
         O     "DB619_State_MPart".Cycle[1].LastStanbyTimeTool;
         O     "DB110_Interf_Program_M1".Bits.MouldNotReleased;
         =     "DB110_Interf_Program_M1".Bits.LastStandbyTimeTool;
END_REGION

REGION Network 6: Interface signals mixinghead 1 mouldcarrier 1
         A     "DB704_MH_Value".MH_Inerting[1].with_output_without_N2;
         =     "DB614_MH_State".InertingMH[1].Inert_Off_Dry_Shot;

         O     "DB123_MH_IO_Signals".MH[1].IN.MH_Manual_Mode;
         O     "DB123_MH_IO_Signals".MH[1].IN.MH_Auto_Mode;
         AN    "DB824_Error_MH_CP".MH_Control[1].FLT_ShotStopped;
         AN    "DB824_Error_MH_CP".CPiston[1].IPS_defect;
         A     "DB619_State_MPart".Operationmode[1].Auto;
         A     "DB619_State_MPart".Operationmode[1].Active;
         =     #Release_Foaming;
   //------------------------------------------------------------------------------
   //  Freigabe zum automatischen Abruf des Schäumzykluses
   //------------------------------------------------------------------------------
   //-----
         O     "DB005_RS<->Extern".MC_Interface[1].Data_from_MC.Shot_preperation;
         O     "DB005_RS<->Extern".MC_Interface[1].Data_from_MC.Shot_release;
         =     #TempReleasInterface;
   //-----
         O     "DB110_Interf_Program_M1".HM_MC_Fault."01";
         =     "DB123_MH_IO_Signals".MH[1].OUT.MH.K_Fault_MC;
         =     "DB005_RS<->Extern".MC_Interface[1].Data_to_MC.Fault;
   //------------------------------------------------------------------------------
   // Programmno. interface in manual mode
   //------------------------------------------------------------------------------
         L     "DB123_MH_IO_Signals".MH[1].IN.MH_Prog_No_MH;
         A     "DB123_MH_IO_Signals".MH[1].IN.MH_Manual_Mode;
         JC    prnr;
         L     0;
   prnr: T     #Temp_ProgNo_MK1_manual;
   //-----
         A     "DB123_MH_IO_Signals".MH[1].IN.MH_Start;
         A     "DB123_MH_IO_Signals".MH[1].IN.MH_Manual_Mode;
         =     #Start_Zyklus;
   //-----
         O(;
         A     "DB005_RS<->Extern".MC_Interface[1].Data_from_MC.Selected;
         A     "DB123_MH_IO_Signals".MH[1].IN.MH_Stop;
         A     "DB123_MH_IO_Signals".MH[1].IN.MH_Auto_Mode;
         );
         O(;
         A     "DB123_MH_IO_Signals".MH[1].IN.MH_Stop;
         A     "DB123_MH_IO_Signals".MH[1].IN.MH_Manual_Mode;
         );
         =     #Temp_Stop;

   //-----
         CALL  "FC112_IF_SP_MC"
         ( IN_InterfaceNo           := 1,
           IN_PositionFIRST         := "DB110_Interf_Program_M1".FIRST,
           IN_PositionSECOND        := "DB110_Interf_Program_M1".SECOND,
           IN_BCDSwitchPrgrNo_MH    := #Temp_ProgNo_MK1_manual,
           IN_MH_Automatic          := "DB123_MH_IO_Signals".MH[1].IN.MH_Auto_Mode,
           IN_MH_Manual             := "DB123_MH_IO_Signals".MH[1].IN.MH_Manual_Mode,
           IN_Start_MH_Panel        := #Start_Zyklus,  //"DB123_MH_IO_Signals".MH[1].IN.MH_Start
           IN_Stop_MH_Panel         := #Temp_Stop,
           IN_ResetFault            := "DB009_Faults".Faults_Reset_FKT_M1,
           IN_ReleaseSWU            := "DB619_State_MPart".SWU[1].SWU_released."01",
           IN_ReleaseMouldcarrier   := #TempReleasInterface,
           IN_PrgNoSwitchDeselected := "DB123_MH_IO_Signals".MH[1].IN.MH_Auto_Mode,
           IN_ReleaseFoaming        := #Release_Foaming,
           IN_ReleaseCycle          := "DB619_State_MPart".Cycle[1].Release,
           IN_OperationModeAuto     := "DB619_State_MPart".Operationmode[1].Auto,
           IN_OperationModeTest     := "DB619_State_MPart".Operationmode[1].Test,
           IN_LampTest              := "DB619_State_MPart".Operationmode[1].Lamptest,
           IN_CycleRunning          := "DB619_State_MPart".ToolMa[1].StationActive,
           IN_ShotRunning           := "DB619_State_MPart".Cycle[1].ShotRuns,
           IN_LastStandbyTimeCycle  := "DB110_Interf_Program_M1".Bits.LastStandbyTimeTool,
           IN_PulseCycleFinished    := "DB619_State_MPart".Cycle[1].Pulse_ToolFinished,
           OUT_Fault_To_MC          := "DB110_Interf_Program_M1".HM_MC_Fault."01",
           OUT_ShotEnd_To_MC        := "DB110_Interf_Program_M1".HM_MC_Shotend."01",
           OUT_H_MH_Panel           := #H_MH_Panel,  // "DB110_Interf_Program_M1".HM_MC_Lamp."01"
           IO_InterfaceActiveFIFO   := "DB110_Interf_Program_M1".Putin_FIFOlist."01",
           IO_Status                := "DB110_Interf_Program_M1".Status_IF[1],
           IO_Fault                 := "DB825_Error_Interface".Interface_MC[1],
           IO_NewFault              := "DB009_Faults".Faultschanging_M1,
           IO_FaultLevel_1          := "DB009_Faults".Faults_FKT_Grp_1_M1,
           IO_FaultLevel_3          := "DB009_Faults".Faults_FKT_Grp_3_M1
         );
   //-----
   //-
   //- General
   //-
         A     #H_MH_Panel;
         O(;
         A     "DB1900_IF_Robots".State_ABB[1].Output.doIRBInHome;
         A     "DB1900_IF_Robots".State_ABB[1].Output.doIRBinAuto;
         A     "DB1900_IF_Robots".State_ABB[1].Output.doCycleOn;
         AN    "DB1900_IF_Robots".State_ABB[1].Output.doSysError;
         AN    "DB619_State_MPart".Cycle[1].running;
         );
         O(;
         A     "DB1900_IF_Robots".State_ABB[1].Output.doIRBInWaitP;
         A     "DB1900_IF_Robots".State_ABB[1].Output.doInWaitPos;
         );
         AN    "DB619_State_MPart".Operationmode[1].Test;
         O     "DB110_Interf_Program_M1".Test_M01.Spare_0_7;
         =     "DB110_Interf_Program_M1".HM_MC_Lamp."01";
   //----------------------------------------------------------------------------------------
   //     Schnittstelle Presse
   //----------------------------------------------------------------------------------------
         AN    #TempReleasInterface;
         R     "DB005_RS<->Extern".MC_Interface[1].Data_to_MC.Shot_end;
   //
         O     "DB110_Interf_Program_M1".Bits.MouldNotReleased;
         O(;
         A     #TempReleasInterface;
         A     "DB110_Interf_Program_M1".HM_MC_Shotend."01";
         );
         S     "DB005_RS<->Extern".MC_Interface[1].Data_to_MC.Shot_end;
   //
         A     "DB005_RS<->Extern".MC_Interface[1].Data_to_MC.Shot_end;
         =     "DB123_MH_IO_Signals".MH[1].OUT.MH.K_ShotEnd_MC;
   //-----
         A     "DB110_Interf_Program_M1".HM_MC_Fault."01";
         =     "DB005_RS<->Extern".MC_Interface[1].Data_to_MC.Fault;
   //
         A     "DB123_MH_IO_Signals".MH[1].IN.MH_Auto_Mode;
         A     "DB619_State_MPart".Operationmode[1].Auto;
         =     "DB005_RS<->Extern".MC_Interface[1].Data_to_MC.Automatic_mode;
   //
         AN    "DB614_MH_State".MH_Status[1].Switch_Service_ON_OFF;
         =     "DB005_RS<->Extern".MC_Interface[1].Data_to_MC.Service_mode;
   //
         A     "DB619_State_MPart".Cycle[1].ShotRuns;
         =     "DB005_RS<->Extern".MC_Interface[1].Data_to_MC.Shot_runs;
   //
         O     "DB1900_IF_Robots".State_ABB[1].Output.doIRBInHome;
         O     "DB1900_IF_Robots".State_ABB[1].Output.doSafetyArea_1;
         =     "DB005_RS<->Extern".MC_Interface[1].Data_to_MC.Robot_out_of_MC;
   //
         A     "DB005_RS<->Extern".MC_Interface[1].Data_from_MC.Com_control;
         =     "DB005_RS<->Extern".MC_Interface[1].Data_to_MC.Com_Control;
   //
         L     "DB005_RS<->Extern".MC_Interface[1].Data_from_MC.Toolcode;
         T     "DB005_RS<->Extern".MC_Interface[1].Data_to_MC.Toolcode;
   //-----
         A     "DB009_Faults".Faults_Reset_FKT_M1;
         R     "DB825_Error_Interface".Interface_MC[1].FLT_Communication;

         L     s5t#5s;
         AN    "DB005_RS<->Extern".MC_Interface[1].Data_from_MC.Com_control;
         SE    "TIM_FRA_WDG1";

         AN    "TIM_FRA_WDG1";
         AN    "DB825_Error_Interface".Interface_MC[1].FLT_Communication;
         CLR;
         S     "DB825_Error_Interface".Interface_MC[1].FLT_Communication;

   // load number to tool alloc
         AN    "DB790_PlantParameter".Bit.ProgrammNofromInterface;
         JC    NoToolNoFromIF01;

         CALL  "FC5_Check_allocAutoMode"
         ( ToolcodeNo := "DB005_RS<->Extern".MC_Interface[1].Data_from_MC.Toolcode,
           ToolAlloc  := "DB940_Tool_alloc_automatic".Alloc_stationTool[1]
         );

   NoToolNoFromIF01:NOP   0;
END_REGION

REGION Network 7: Interface signals mixinghead 2 mouldcarrier 2
         A     "DB704_MH_Value".MH_Inerting[1].with_output_without_N2;
         =     "DB614_MH_State".InertingMH[1].Inert_Off_Dry_Shot;

         O     "DB123_MH_IO_Signals".MH[1].IN.MH_Manual_Mode;
         O     "DB123_MH_IO_Signals".MH[1].IN.MH_Auto_Mode;
         AN    "DB824_Error_MH_CP".MH_Control[1].FLT_ShotStopped;
         AN    "DB824_Error_MH_CP".CPiston[1].IPS_defect;
         A     "DB619_State_MPart".Operationmode[1].Auto;
         A     "DB619_State_MPart".Operationmode[1].Active;
         =     #Release_Foaming;
   //------------------------------------------------------------------------------
   //  Freigabe zum automatischen Abruf des Schäumzykluses
   //------------------------------------------------------------------------------
   //-----
         O     "DB005_RS<->Extern".MC_Interface[2].Data_from_MC.Shot_preperation;
         O     "DB005_RS<->Extern".MC_Interface[2].Data_from_MC.Shot_release;
         =     #TempReleasInterface;
   //-----
         O     "DB110_Interf_Program_M1".HM_MC_Fault."02";
         =     "DB005_RS<->Extern".MC_Interface[2].Data_to_MC.Fault;
   //-----
         A     "DB123_MH_IO_Signals".MH[1].IN.MH_Start;
         A     "DB123_MH_IO_Signals".MH[1].IN.MH_Manual_Mode;
         =     #Start_Zyklus;
   //-----
         A     "DB005_RS<->Extern".MC_Interface[2].Data_from_MC.Selected;
         A     "DB123_MH_IO_Signals".MH[1].IN.MH_Stop;
         =     #Temp_Stop;
   //-----
         CALL  "FC112_IF_SP_MC"
         ( IN_InterfaceNo           := 2,
           IN_PositionFIRST         := "DB110_Interf_Program_M1".FIRST,
           IN_PositionSECOND        := "DB110_Interf_Program_M1".SECOND,
           IN_BCDSwitchPrgrNo_MH    := 0,
           IN_MH_Automatic          := "DB123_MH_IO_Signals".MH[1].IN.MH_Auto_Mode,
           IN_MH_Manual             := false,
           IN_Start_MH_Panel        := #Start_Zyklus,
           IN_Stop_MH_Panel         := #Temp_Stop,
           IN_ResetFault            := "DB009_Faults".Faults_Reset_FKT_M1,
           IN_ReleaseSWU            := "DB619_State_MPart".SWU[1].SWU_released."01",
           IN_ReleaseMouldcarrier   := #TempReleasInterface,
           IN_PrgNoSwitchDeselected := "DB123_MH_IO_Signals".MH[1].IN.MH_Auto_Mode,
           IN_ReleaseFoaming        := #Release_Foaming,
           IN_ReleaseCycle          := "DB619_State_MPart".Cycle[1].Release,
           IN_OperationModeAuto     := "DB619_State_MPart".Operationmode[1].Auto,
           IN_OperationModeTest     := "DB619_State_MPart".Operationmode[1].Test,
           IN_LampTest              := "DB619_State_MPart".Operationmode[1].Lamptest,
           IN_CycleRunning          := "DB619_State_MPart".ToolMa[1].StationActive,
           IN_ShotRunning           := "DB619_State_MPart".Cycle[1].ShotRuns,
           IN_LastStandbyTimeCycle  := "DB110_Interf_Program_M1".Bits.LastStandbyTimeTool,
           IN_PulseCycleFinished    := "DB619_State_MPart".Cycle[1].Pulse_ToolFinished,
           OUT_Fault_To_MC          := "DB110_Interf_Program_M1".HM_MC_Fault."02",
           OUT_ShotEnd_To_MC        := "DB110_Interf_Program_M1".HM_MC_Shotend."02",
           OUT_H_MH_Panel           := #H_MH_Panel,  // "DB110_Interf_Program_M1".HM_MC_Lamp."02"
           IO_InterfaceActiveFIFO   := "DB110_Interf_Program_M1".Putin_FIFOlist."02",
           IO_Status                := "DB110_Interf_Program_M1".Status_IF[2],
           IO_Fault                 := "DB825_Error_Interface".Interface_MC[2],
           IO_NewFault              := "DB009_Faults".Faultschanging_M1,
           IO_FaultLevel_1          := "DB009_Faults".Faults_FKT_Grp_1_M1,
           IO_FaultLevel_3          := "DB009_Faults".Faults_FKT_Grp_3_M1
         );
   //-----
   //-
   //- General
   //-
         A     #H_MH_Panel;
         O(;
         A     "DB1900_IF_Robots".State_ABB[1].Output.doIRBInHome;
         A     "DB1900_IF_Robots".State_ABB[1].Output.doIRBinAuto;
         A     "DB1900_IF_Robots".State_ABB[1].Output.doCycleOn;
         AN    "DB1900_IF_Robots".State_ABB[1].Output.doSysError;
         AN    "DB619_State_MPart".Cycle[1].running;
         );
         O(;
         A     "DB1900_IF_Robots".State_ABB[1].Output.doIRBInWaitP;
         A     "DB1900_IF_Robots".State_ABB[1].Output.doInWaitPos;
         );
         =     "DB110_Interf_Program_M1".HM_MC_Lamp."02";
   //----------------------------------------------------------------------------------------
   //     Schnittstelle Presse
   //----------------------------------------------------------------------------------------
         AN    #TempReleasInterface;
         R     "DB005_RS<->Extern".MC_Interface[2].Data_to_MC.Shot_end;
   //
         O     "DB110_Interf_Program_M1".Bits.MouldNotReleased;
         O(;
         A     #TempReleasInterface;
         A     "DB110_Interf_Program_M1".HM_MC_Shotend."02";
         );
         S     "DB005_RS<->Extern".MC_Interface[2].Data_to_MC.Shot_end;
   //-----
         A     "DB110_Interf_Program_M1".HM_MC_Fault."02";
         =     "DB005_RS<->Extern".MC_Interface[2].Data_to_MC.Fault;
   //
         A     "DB123_MH_IO_Signals".MH[1].IN.MH_Auto_Mode;
         A     "DB619_State_MPart".Operationmode[1].Auto;
         =     "DB005_RS<->Extern".MC_Interface[2].Data_to_MC.Automatic_mode;
   //
         AN    "DB614_MH_State".MH_Status[1].Switch_Service_ON_OFF;
         =     "DB005_RS<->Extern".MC_Interface[2].Data_to_MC.Service_mode;
   //
         A     "DB619_State_MPart".Cycle[1].ShotRuns;
         =     "DB005_RS<->Extern".MC_Interface[2].Data_to_MC.Shot_runs;
   //
         O     "DB1900_IF_Robots".State_ABB[1].Output.doIRBInHome;
         O     "DB1900_IF_Robots".State_ABB[1].Output.doSafetyArea_2;
         =     "DB005_RS<->Extern".MC_Interface[2].Data_to_MC.Robot_out_of_MC;
   //
         A     "DB005_RS<->Extern".MC_Interface[2].Data_from_MC.Com_control;
         =     "DB005_RS<->Extern".MC_Interface[2].Data_to_MC.Com_Control;
   //
         L     "DB005_RS<->Extern".MC_Interface[2].Data_from_MC.Toolcode;
         T     "DB005_RS<->Extern".MC_Interface[2].Data_to_MC.Toolcode;
   //-----
         A     "DB009_Faults".Faults_Reset_FKT_M1;
         R     "DB825_Error_Interface".Interface_MC[2].FLT_Communication;

         L     s5t#5s;
         AN    "DB005_RS<->Extern".MC_Interface[2].Data_from_MC.Com_control;
         SE    "TIM_FRA_WDG2";

         AN    "TIM_FRA_WDG2";
         AN    "DB825_Error_Interface".Interface_MC[2].FLT_Communication;
         CLR;
         S     "DB825_Error_Interface".Interface_MC[2].FLT_Communication;

   // load number to tool alloc
         AN    "DB790_PlantParameter".Bit.ProgrammNofromInterface;
         JC    NoToolNoFromIF02;

         CALL  "FC5_Check_allocAutoMode"
         ( ToolcodeNo := "DB005_RS<->Extern".MC_Interface[2].Data_from_MC.Toolcode,
           ToolAlloc  := "DB940_Tool_alloc_automatic".Alloc_stationTool[2]
         );

   NoToolNoFromIF02:NOP   0;
END_REGION

REGION Network 8: Interface signals mixinghead 3 mouldcarrier 3
         A     "DB704_MH_Value".MH_Inerting[1].with_output_without_N2;
         =     "DB614_MH_State".InertingMH[1].Inert_Off_Dry_Shot;

         O     "DB123_MH_IO_Signals".MH[1].IN.MH_Manual_Mode;
         O     "DB123_MH_IO_Signals".MH[1].IN.MH_Auto_Mode;
         AN    "DB824_Error_MH_CP".MH_Control[1].FLT_ShotStopped;
         AN    "DB824_Error_MH_CP".CPiston[1].IPS_defect;
         A     "DB619_State_MPart".Operationmode[1].Auto;
         A     "DB619_State_MPart".Operationmode[1].Active;
         =     #Release_Foaming;
   //------------------------------------------------------------------------------
   //  Freigabe zum automatischen Abruf des Schäumzykluses
   //------------------------------------------------------------------------------
   //-----
         O     "DB005_RS<->Extern".MC_Interface[3].Data_from_MC.Shot_preperation;
         O     "DB005_RS<->Extern".MC_Interface[3].Data_from_MC.Shot_release;
         =     #TempReleasInterface;
   //-----
         O     "DB110_Interf_Program_M1".HM_MC_Fault."03";
         =     "DB005_RS<->Extern".MC_Interface[3].Data_to_MC.Fault;
   //-----
         A     "DB123_MH_IO_Signals".MH[1].IN.MH_Start;
         A     "DB123_MH_IO_Signals".MH[1].IN.MH_Manual_Mode;
         =     #Start_Zyklus;
   //-----
         A     "DB005_RS<->Extern".MC_Interface[3].Data_from_MC.Selected;
         A     "DB123_MH_IO_Signals".MH[1].IN.MH_Stop;
         =     #Temp_Stop;
   //-----
         CALL  "FC112_IF_SP_MC"
         ( IN_InterfaceNo           := 3,
           IN_PositionFIRST         := "DB110_Interf_Program_M1".FIRST,
           IN_PositionSECOND        := "DB110_Interf_Program_M1".SECOND,
           IN_BCDSwitchPrgrNo_MH    := 0,
           IN_MH_Automatic          := "DB123_MH_IO_Signals".MH[1].IN.MH_Auto_Mode,
           IN_MH_Manual             := false,
           IN_Start_MH_Panel        := #Start_Zyklus,
           IN_Stop_MH_Panel         := #Temp_Stop,
           IN_ResetFault            := "DB009_Faults".Faults_Reset_FKT_M1,
           IN_ReleaseSWU            := "DB619_State_MPart".SWU[1].SWU_released."01",
           IN_ReleaseMouldcarrier   := #TempReleasInterface,
           IN_PrgNoSwitchDeselected := "DB123_MH_IO_Signals".MH[1].IN.MH_Auto_Mode,
           IN_ReleaseFoaming        := #Release_Foaming,
           IN_ReleaseCycle          := "DB619_State_MPart".Cycle[1].Release,
           IN_OperationModeAuto     := "DB619_State_MPart".Operationmode[1].Auto,
           IN_OperationModeTest     := "DB619_State_MPart".Operationmode[1].Test,
           IN_LampTest              := "DB619_State_MPart".Operationmode[1].Lamptest,
           IN_CycleRunning          := "DB619_State_MPart".ToolMa[1].StationActive,
           IN_ShotRunning           := "DB619_State_MPart".Cycle[1].ShotRuns,
           IN_LastStandbyTimeCycle  := "DB110_Interf_Program_M1".Bits.LastStandbyTimeTool,
           IN_PulseCycleFinished    := "DB619_State_MPart".Cycle[1].Pulse_ToolFinished,
           OUT_Fault_To_MC          := "DB110_Interf_Program_M1".HM_MC_Fault."03",
           OUT_ShotEnd_To_MC        := "DB110_Interf_Program_M1".HM_MC_Shotend."03",
           OUT_H_MH_Panel           := #H_MH_Panel,  // "DB110_Interf_Program_M1".HM_MC_Lamp."03"
           IO_InterfaceActiveFIFO   := "DB110_Interf_Program_M1".Putin_FIFOlist."03",
           IO_Status                := "DB110_Interf_Program_M1".Status_IF[3],
           IO_Fault                 := "DB825_Error_Interface".Interface_MC[3],
           IO_NewFault              := "DB009_Faults".Faultschanging_M1,
           IO_FaultLevel_1          := "DB009_Faults".Faults_FKT_Grp_1_M1,
           IO_FaultLevel_3          := "DB009_Faults".Faults_FKT_Grp_3_M1
         );
   //-----
   //-
   //- General
   //-
         A     #H_MH_Panel;
         O(;
         A     "DB1900_IF_Robots".State_ABB[1].Output.doIRBInHome;
         A     "DB1900_IF_Robots".State_ABB[1].Output.doIRBinAuto;
         A     "DB1900_IF_Robots".State_ABB[1].Output.doCycleOn;
         AN    "DB1900_IF_Robots".State_ABB[1].Output.doSysError;
         AN    "DB619_State_MPart".Cycle[1].running;
         );
         O(;
         A     "DB1900_IF_Robots".State_ABB[1].Output.doIRBInWaitP;
         A     "DB1900_IF_Robots".State_ABB[1].Output.doInWaitPos;
         );
         =     "DB110_Interf_Program_M1".HM_MC_Lamp."03";
   //----------------------------------------------------------------------------------------
   //     Schnittstelle Presse
   //----------------------------------------------------------------------------------------
         AN    #TempReleasInterface;
         R     "DB005_RS<->Extern".MC_Interface[3].Data_to_MC.Shot_end;
   //
         O     "DB110_Interf_Program_M1".Bits.MouldNotReleased;
         O(;
         A     #TempReleasInterface;
         A     "DB110_Interf_Program_M1".HM_MC_Shotend."03";
         );
         S     "DB005_RS<->Extern".MC_Interface[3].Data_to_MC.Shot_end;
   //-----
         A     "DB110_Interf_Program_M1".HM_MC_Fault."03";
         =     "DB005_RS<->Extern".MC_Interface[3].Data_to_MC.Fault;
   //
         A     "DB123_MH_IO_Signals".MH[1].IN.MH_Auto_Mode;
         A     "DB619_State_MPart".Operationmode[1].Auto;
         =     "DB005_RS<->Extern".MC_Interface[3].Data_to_MC.Automatic_mode;
   //
         AN    "DB614_MH_State".MH_Status[1].Switch_Service_ON_OFF;
         =     "DB005_RS<->Extern".MC_Interface[3].Data_to_MC.Service_mode;
   //
         A     "DB619_State_MPart".Cycle[1].ShotRuns;
         =     "DB005_RS<->Extern".MC_Interface[3].Data_to_MC.Shot_runs;
   //
         O     "DB1900_IF_Robots".State_ABB[1].Output.doIRBInHome;
         O     "DB1900_IF_Robots".State_ABB[1].Output.doSafetyArea_3;
         =     "DB005_RS<->Extern".MC_Interface[3].Data_to_MC.Robot_out_of_MC;
   //
         A     "DB005_RS<->Extern".MC_Interface[3].Data_from_MC.Com_control;
         =     "DB005_RS<->Extern".MC_Interface[3].Data_to_MC.Com_Control;
   //
         L     "DB005_RS<->Extern".MC_Interface[3].Data_from_MC.Toolcode;
         T     "DB005_RS<->Extern".MC_Interface[3].Data_to_MC.Toolcode;
   //-----
         A     "DB009_Faults".Faults_Reset_FKT_M1;
         R     "DB825_Error_Interface".Interface_MC[3].FLT_Communication;

         L     s5t#5s;
         AN    "DB005_RS<->Extern".MC_Interface[3].Data_from_MC.Com_control;
         SE    "TIM_FRA_WDG3";

         AN    "TIM_FRA_WDG3";
         A     "With_MC03";
         AN    "DB825_Error_Interface".Interface_MC[3].FLT_Communication;
         S     "DB825_Error_Interface".Interface_MC[3].FLT_Communication;

   // load number to tool alloc
         AN    "DB790_PlantParameter".Bit.ProgrammNofromInterface;
         JC    NoToolNoFromIF03;

         CALL  "FC5_Check_allocAutoMode"
         ( ToolcodeNo := "DB005_RS<->Extern".MC_Interface[3].Data_from_MC.Toolcode,
           ToolAlloc  := "DB940_Tool_alloc_automatic".Alloc_stationTool[3]
         );

   NoToolNoFromIF03:NOP   0;
END_REGION

REGION Network 9: Interface signals mixinghead 4 mouldcarrier 4
         A     "DB704_MH_Value".MH_Inerting[1].with_output_without_N2;
         =     "DB614_MH_State".InertingMH[1].Inert_Off_Dry_Shot;

         O     "DB123_MH_IO_Signals".MH[1].IN.MH_Manual_Mode;
         O     "DB123_MH_IO_Signals".MH[1].IN.MH_Auto_Mode;
         AN    "DB824_Error_MH_CP".MH_Control[1].FLT_ShotStopped;
         AN    "DB824_Error_MH_CP".CPiston[1].IPS_defect;
         A     "DB619_State_MPart".Operationmode[1].Auto;
         A     "DB619_State_MPart".Operationmode[1].Active;
         =     #Release_Foaming;
   //------------------------------------------------------------------------------
   //  Freigabe zum automatischen Abruf des Schäumzykluses
   //------------------------------------------------------------------------------
   //-----
         O     "DB005_RS<->Extern".MC_Interface[4].Data_from_MC.Shot_preperation;
         O     "DB005_RS<->Extern".MC_Interface[4].Data_from_MC.Shot_release;
         =     #TempReleasInterface;
   //-----
         O     "DB110_Interf_Program_M1".HM_MC_Fault."04";
         =     "DB005_RS<->Extern".MC_Interface[4].Data_to_MC.Fault;
   //-----
         A     "DB123_MH_IO_Signals".MH[1].IN.MH_Start;
         A     "DB123_MH_IO_Signals".MH[1].IN.MH_Manual_Mode;
         =     #Start_Zyklus;
   //-----
         A     "DB005_RS<->Extern".MC_Interface[4].Data_from_MC.Selected;
         A     "DB123_MH_IO_Signals".MH[1].IN.MH_Stop;
         =     #Temp_Stop;
   //-----
         CALL  "FC112_IF_SP_MC"
         ( IN_InterfaceNo           := 4,
           IN_PositionFIRST         := "DB110_Interf_Program_M1".FIRST,
           IN_PositionSECOND        := "DB110_Interf_Program_M1".SECOND,
           IN_BCDSwitchPrgrNo_MH    := 0,
           IN_MH_Automatic          := "DB123_MH_IO_Signals".MH[1].IN.MH_Auto_Mode,
           IN_MH_Manual             := false,
           IN_Start_MH_Panel        := #Start_Zyklus,
           IN_Stop_MH_Panel         := #Temp_Stop,
           IN_ResetFault            := "DB009_Faults".Faults_Reset_FKT_M1,
           IN_ReleaseSWU            := "DB619_State_MPart".SWU[1].SWU_released."01",
           IN_ReleaseMouldcarrier   := #TempReleasInterface,
           IN_PrgNoSwitchDeselected := "DB123_MH_IO_Signals".MH[1].IN.MH_Auto_Mode,
           IN_ReleaseFoaming        := #Release_Foaming,
           IN_ReleaseCycle          := "DB619_State_MPart".Cycle[1].Release,
           IN_OperationModeAuto     := "DB619_State_MPart".Operationmode[1].Auto,
           IN_OperationModeTest     := "DB619_State_MPart".Operationmode[1].Test,
           IN_LampTest              := "DB619_State_MPart".Operationmode[1].Lamptest,
           IN_CycleRunning          := "DB619_State_MPart".ToolMa[1].StationActive,
           IN_ShotRunning           := "DB619_State_MPart".Cycle[1].ShotRuns,
           IN_LastStandbyTimeCycle  := "DB110_Interf_Program_M1".Bits.LastStandbyTimeTool,
           IN_PulseCycleFinished    := "DB619_State_MPart".Cycle[1].Pulse_ToolFinished,
           OUT_Fault_To_MC          := "DB110_Interf_Program_M1".HM_MC_Fault."04",
           OUT_ShotEnd_To_MC        := "DB110_Interf_Program_M1".HM_MC_Shotend."04",
           OUT_H_MH_Panel           := #H_MH_Panel,  // "DB110_Interf_Program_M1".HM_MC_Lamp."04"
           IO_InterfaceActiveFIFO   := "DB110_Interf_Program_M1".Putin_FIFOlist."04",
           IO_Status                := "DB110_Interf_Program_M1".Status_IF[4],
           IO_Fault                 := "DB825_Error_Interface".Interface_MC[4],
           IO_NewFault              := "DB009_Faults".Faultschanging_M1,
           IO_FaultLevel_1          := "DB009_Faults".Faults_FKT_Grp_1_M1,
           IO_FaultLevel_3          := "DB009_Faults".Faults_FKT_Grp_3_M1
         );
   //-----
   //-
   //- General
   //-
         A     #H_MH_Panel;
         O(;
         A     "DB1900_IF_Robots".State_ABB[1].Output.doIRBInHome;
         A     "DB1900_IF_Robots".State_ABB[1].Output.doIRBinAuto;
         A     "DB1900_IF_Robots".State_ABB[1].Output.doCycleOn;
         AN    "DB1900_IF_Robots".State_ABB[1].Output.doSysError;
         AN    "DB619_State_MPart".Cycle[1].running;
         );
         O(;
         A     "DB1900_IF_Robots".State_ABB[1].Output.doIRBInWaitP;
         A     "DB1900_IF_Robots".State_ABB[1].Output.doInWaitPos;
         );
         =     "DB110_Interf_Program_M1".HM_MC_Lamp."04";
   //----------------------------------------------------------------------------------------
   //     Schnittstelle Presse
   //----------------------------------------------------------------------------------------
         AN    #TempReleasInterface;
         R     "DB005_RS<->Extern".MC_Interface[4].Data_to_MC.Shot_end;
   //
         O     "DB110_Interf_Program_M1".Bits.MouldNotReleased;
         O(;
         A     #TempReleasInterface;
         A     "DB110_Interf_Program_M1".HM_MC_Shotend."04";
         );
         S     "DB005_RS<->Extern".MC_Interface[4].Data_to_MC.Shot_end;
   //-----
         A     "DB110_Interf_Program_M1".HM_MC_Fault."04";
         =     "DB005_RS<->Extern".MC_Interface[4].Data_to_MC.Fault;
   //
         A     "DB123_MH_IO_Signals".MH[1].IN.MH_Auto_Mode;
         A     "DB619_State_MPart".Operationmode[1].Auto;
         =     "DB005_RS<->Extern".MC_Interface[4].Data_to_MC.Automatic_mode;
   //
         AN    "DB614_MH_State".MH_Status[1].Switch_Service_ON_OFF;
         =     "DB005_RS<->Extern".MC_Interface[4].Data_to_MC.Service_mode;
   //
         A     "DB619_State_MPart".Cycle[1].ShotRuns;
         =     "DB005_RS<->Extern".MC_Interface[4].Data_to_MC.Shot_runs;
   //
         O     "DB1900_IF_Robots".State_ABB[1].Output.doIRBInHome;
         O     "DB1900_IF_Robots".State_ABB[1].Output.doSafetyArea_4;
         =     "DB005_RS<->Extern".MC_Interface[4].Data_to_MC.Robot_out_of_MC;
   //
         A     "DB005_RS<->Extern".MC_Interface[4].Data_from_MC.Com_control;
         =     "DB005_RS<->Extern".MC_Interface[4].Data_to_MC.Com_Control;
   //
         L     "DB005_RS<->Extern".MC_Interface[4].Data_from_MC.Toolcode;
         T     "DB005_RS<->Extern".MC_Interface[4].Data_to_MC.Toolcode;
   //-----
         A     "DB009_Faults".Faults_Reset_FKT_M1;
         R     "DB825_Error_Interface".Interface_MC[4].FLT_Communication;

         L     s5t#5s;
         AN    "DB005_RS<->Extern".MC_Interface[4].Data_from_MC.Com_control;
         SE    "TIM_FRA_WDG4";

         AN    "TIM_FRA_WDG4";
         A     "With_MC04";
         AN    "DB825_Error_Interface".Interface_MC[4].FLT_Communication;
         S     "DB825_Error_Interface".Interface_MC[4].FLT_Communication;

   // load number to tool alloc
         AN    "DB790_PlantParameter".Bit.ProgrammNofromInterface;
         JC    NoToolNoFromIF04;

         CALL  "FC5_Check_allocAutoMode"
         ( ToolcodeNo := "DB005_RS<->Extern".MC_Interface[4].Data_from_MC.Toolcode,
           ToolAlloc  := "DB940_Tool_alloc_automatic".Alloc_stationTool[4]
         );

   NoToolNoFromIF04:NOP   0;
END_REGION

REGION Network 10: Test with test valves
   //     CALL  "FC115_Testen"
   //         IN_Betriebsart_Testen   :="DB619_State_MPart".Operationmode[1].Test
   //         IN_Betriebsart_Betrieb  :="DB619_State_MPart".Operationmode[1].Operation
   //         IN_Lampentest           :="DB619_State_MPart".Operationmode[1].Lamptest
   //         IN_Start_Testen_K1      :="T_Start_Test_C1"
   //         IN_Start_Testen_K2      :="T_Start_Test_C2"
   //         IN_Start_Testen_K3      :=FALSE
   //         IN_Start_Testen_K4      :=FALSE
   //         IN_Stop_Testen          :="T_Stop_Test"
   //         IN_Stoerung_Gruppe_1    :="DB009_Faults".Faults_FKT_Grp_1_M1
   //         IN_Zyklus_Freigabe      :="DB619_State_MPart".Cycle[1].Release
   //         IN_Zyklus_laeuft        :="DB619_State_MPart".ToolMa[1].StationActive
   //         IN_Zyklus_Schuss_laeuft :="DB619_State_MPart".Cycle[1].ShotRuns
   //         IN_Imp_Zyklus_Ende      :="DB619_State_MPart".Cycle[1].Pulse_ToolFinished
   //         IN_Zyklus_KLZ2_u_ff     :="DB619_State_MPart".Cycle[1].LastStanbyTimeTool
   //         OUT_H_Testen_K1         :="H_Test_C1"
   //         OUT_H_Testen_K2         :="H_Test_C2"
   //         OUT_H_Testen_K3         :=#Dummy
   //         OUT_H_Testen_K4         :=#Dummy
   //         OUT_V_Testen_K1         :="V_Test_C1"
   //         OUT_V_Testen_K2         :="V_Test_C2"
   //         OUT_V_Testen_K3         :=#Dummy
   //         OUT_V_Testen_K4         :=#Dummy
   //         IO_Status               :="DB110_Interf_Program_M1".Test_M01
   //
END_REGION

REGION Network 11: LED mixing head panel
   //-----
         A     "DB110_Interf_Program_M1".HM_MC_Lamp."01";
         O;
         A     "DB110_Interf_Program_M1".Status_IF[2].IF_is_on_1_Position;
         A     "DB110_Interf_Program_M1".HM_MC_Lamp."02";
         O;
         A     "DB110_Interf_Program_M1".Status_IF[3].IF_is_on_1_Position;
         A     "DB110_Interf_Program_M1".HM_MC_Lamp."03";
         O;
         A     "DB110_Interf_Program_M1".Status_IF[4].IF_is_on_1_Position;
         A     "DB110_Interf_Program_M1".HM_MC_Lamp."04";
         O;
         A     "DB110_Interf_Program_M1".Status_IF[5].IF_is_on_1_Position;
         A     "DB110_Interf_Program_M1".HM_MC_Lamp."05";
         =     "DB123_MH_IO_Signals".MH[1].OUT.MH.H_Rel_Foaming_MH;
END_REGION

REGION Network 12: Start cycle
         A     "DB1900_IF_Robots".State_Robots[1].ReadyForStartCycle;
         A     "DB123_MH_IO_Signals".MH[1].IN.MH_Auto_Mode;
         O     "DB123_MH_IO_Signals".MH[1].IN.MH_Manual_Mode;
         A(;
         O     "DB110_Interf_Program_M1".Status_IF[1].Start_to_Cycle;
         O     "DB110_Interf_Program_M1".Status_IF[2].Start_to_Cycle;
         O     "DB110_Interf_Program_M1".Status_IF[3].Start_to_Cycle;
         O     "DB110_Interf_Program_M1".Status_IF[4].Start_to_Cycle;
         O     "DB110_Interf_Program_M1".Status_IF[5].Start_to_Cycle;
         O     "DB110_Interf_Program_M1".Status_IF[6].Start_to_Cycle;
         O     "DB110_Interf_Program_M1".Status_IF[7].Start_to_Cycle;
         O     "DB110_Interf_Program_M1".Status_IF[8].Start_to_Cycle;
         O     "DB110_Interf_Program_M1".Status_IF[9].Start_to_Cycle;
         O     "DB110_Interf_Program_M1".Status_IF[10].Start_to_Cycle;
         );
         O     "DB110_Interf_Program_M1".Test_M01.Start_to_Cycle;
         =     #Start_Zyklus;
END_REGION

REGION Network 13: Stop cycle
         O     "DB110_Interf_Program_M1".Status_IF[1].Stop_to_Cycle;
         O     "DB110_Interf_Program_M1".Status_IF[2].Stop_to_Cycle;
         O     "DB110_Interf_Program_M1".Status_IF[3].Stop_to_Cycle;
         O     "DB110_Interf_Program_M1".Status_IF[4].Stop_to_Cycle;
         O     "DB110_Interf_Program_M1".Status_IF[5].Stop_to_Cycle;
         O     "DB110_Interf_Program_M1".Status_IF[6].Stop_to_Cycle;
         O     "DB110_Interf_Program_M1".Status_IF[7].Stop_to_Cycle;
         O     "DB110_Interf_Program_M1".Status_IF[8].Stop_to_Cycle;
         O     "DB110_Interf_Program_M1".Status_IF[9].Stop_to_Cycle;
         O     "DB110_Interf_Program_M1".Status_IF[10].Stop_to_Cycle;
         O     "DB110_Interf_Program_M1".Test_M01.Stop_to_Cycle;
         =     "DB110_Interf_Program_M1".Bits.Stop_Cycle;
         =     "DB619_State_MPart".ToolMa[1].StopCycle;
END_REGION

REGION Network 14: Station number (Program number) to select mould no. ->FB930
         A     #Start_Zyklus;
         AN    "DB619_State_MPart".ToolMa[1].StopCycle;
         JCN   GOON;
   ///----------
         A     "DB619_State_MPart".Operationmode[1].Test;
         JC    Test;
   ///----------
         AN    "DB110_Interf_Program_M1".Status_IF[1].IF_is_on_1_Position;
         JC    SS_2;
   ///----------
         A     "DB123_MH_IO_Signals".MH[1].IN.MH_Auto_Mode;
         JC    SS1A;
   ///----------
         L     #Temp_ProgNo_MK1_manual;
         L     "DB704_MH_Value".Mixinghead[1].pRrgNumberManual;
         +I;
         T     "DB110_Interf_Program_M1".Program_No_01;
         JU    ENDE;
   ///----------
   SS1A: NOP   0;
         AN    "DB005_RS<->Extern".MC_Interface[1].Data_from_MC.Shot_preperation;
         AN    "DB005_RS<->Extern".MC_Interface[1].Data_from_MC.Shot_release;
         ON    "DB619_State_MPart".SWU[1].SWU_released."01";
         JC    ENDE;
   ///----------
         L     1;
         T     "DB110_Interf_Program_M1".Program_No_01;

         L     1;
         T     "DB110_Interf_Program_M1".MixingHeadNo;
         T     "DB110_Interf_Program_M1".Robot_01.MC_Place_Number;

         L     "DB005_RS<->Extern".MC_Interface[1].Data_from_MC.Angle_frame_foaming_pos;
         L     7.0;
         <=R;
         L     1;  //      L     "DB005_RS<->Extern".MC_Interface[1].Data_from_MC.Toolcode
         JC    ProRob01;
         L     1;  // L     "DB005_RS<->Extern".MC_Interface[1].Data_from_MC.Toolcode
         L     100;
         +I;
   ProRob01:T     "DB110_Interf_Program_M1".Robot_01.Robot_ProgNo_Mould_1;
         JU    ENDE;
   ///----------
   SS_2: NOP   0;
         AN    "DB110_Interf_Program_M1".Status_IF[2].IF_is_on_1_Position;
         JC    SS_3;
         A     "DB123_MH_IO_Signals".MH[1].IN.MH_Auto_Mode;
         JC    SS2A;
   ///----------
         L     0;
         T     "DB110_Interf_Program_M1".Program_No_01;
         JU    ENDE;
   ///----------
   SS2A: NOP   0;
         AN    "DB005_RS<->Extern".MC_Interface[2].Data_from_MC.Shot_preperation;
         AN    "DB005_RS<->Extern".MC_Interface[2].Data_from_MC.Shot_release;
         ON    "DB619_State_MPart".SWU[1].SWU_released."01";
         JC    ENDE;
   ///----------
         L     2;
         T     "DB110_Interf_Program_M1".Program_No_01;

         L     1;
         T     "DB110_Interf_Program_M1".MixingHeadNo;

         L     2;
         T     "DB110_Interf_Program_M1".Robot_01.MC_Place_Number;

         L     "DB005_RS<->Extern".MC_Interface[2].Data_from_MC.Angle_frame_foaming_pos;
         L     7.0;
         <=R;
         L     "DB005_RS<->Extern".MC_Interface[2].Data_from_MC.Toolcode;
         JC    ProRob02;
         L     "DB005_RS<->Extern".MC_Interface[2].Data_from_MC.Toolcode;
         L     100;
         +I;
   ProRob02:T     "DB110_Interf_Program_M1".Robot_01.Robot_ProgNo_Mould_1;

   ///----------
   SS_3: NOP   0;
         AN    "DB110_Interf_Program_M1".Status_IF[3].IF_is_on_1_Position;
         JC    SS_4;
         A     "DB123_MH_IO_Signals".MH[1].IN.MH_Auto_Mode;
         JC    SS3A;
   ///----------
         L     0;
         T     "DB110_Interf_Program_M1".Program_No_01;
         JU    ENDE;
   ///----------
   SS3A: NOP   0;
         AN    "DB005_RS<->Extern".MC_Interface[3].Data_from_MC.Shot_preperation;
         AN    "DB005_RS<->Extern".MC_Interface[3].Data_from_MC.Shot_release;
         ON    "DB619_State_MPart".SWU[1].SWU_released."01";
         JC    ENDE;
   ///----------
         L     3;
         T     "DB110_Interf_Program_M1".Program_No_01;

         L     1;
         T     "DB110_Interf_Program_M1".MixingHeadNo;

         L     3;
         T     "DB110_Interf_Program_M1".Robot_01.MC_Place_Number;

         L     "DB005_RS<->Extern".MC_Interface[3].Data_from_MC.Angle_frame_foaming_pos;
         L     7.0;
         <=R;
         L     "DB005_RS<->Extern".MC_Interface[3].Data_from_MC.Toolcode;
         JC    ProRob03;
         L     "DB005_RS<->Extern".MC_Interface[3].Data_from_MC.Toolcode;
         L     100;
         +I;
   ProRob03:T     "DB110_Interf_Program_M1".Robot_01.Robot_ProgNo_Mould_1;
         JU    ENDE;

   ///----------
   SS_4: NOP   0;
         AN    "DB110_Interf_Program_M1".Status_IF[4].IF_is_on_1_Position;
         JC    SS_5;
         A     "DB123_MH_IO_Signals".MH[1].IN.MH_Auto_Mode;
         JC    SS4A;
   ///----------
         L     0;
         T     "DB110_Interf_Program_M1".Program_No_01;
         JU    ENDE;
   ///----------
   SS4A: NOP   0;
         AN    "DB005_RS<->Extern".MC_Interface[4].Data_from_MC.Shot_preperation;
         AN    "DB005_RS<->Extern".MC_Interface[4].Data_from_MC.Shot_release;
         ON    "DB619_State_MPart".SWU[1].SWU_released."01";
         JC    ENDE;
   ///----------
         L     4;
         T     "DB110_Interf_Program_M1".Program_No_01;

         L     1;
         T     "DB110_Interf_Program_M1".MixingHeadNo;

         L     4;
         T     "DB110_Interf_Program_M1".Robot_01.MC_Place_Number;

         L     "DB005_RS<->Extern".MC_Interface[4].Data_from_MC.Angle_frame_foaming_pos;
         L     7.0;
         <=R;
         L     "DB005_RS<->Extern".MC_Interface[4].Data_from_MC.Toolcode;
         JC    ProRob04;
         L     "DB005_RS<->Extern".MC_Interface[4].Data_from_MC.Toolcode;
         L     100;
         +I;
   ProRob04:T     "DB110_Interf_Program_M1".Robot_01.Robot_ProgNo_Mould_1;
         JU    ENDE;
   ///----------
   SS_5: NOP   0;
         AN    "DB110_Interf_Program_M1".Status_IF[5].IF_is_on_1_Position;
         JC    SS_6;
         A     "DB123_MH_IO_Signals".MH[1].IN.MH_Auto_Mode;
         JC    SS5A;
   ///----------
         L     0;
         T     "DB110_Interf_Program_M1".Program_No_01;
         JU    ENDE;
   ///----------
   SS5A: NOP   0;
         AN    "DB005_RS<->Extern".MC_Interface[5].Data_from_MC.Shot_preperation;
         AN    "DB005_RS<->Extern".MC_Interface[5].Data_from_MC.Shot_release;
         ON    "DB619_State_MPart".SWU[1].SWU_released."01";
         JC    ENDE;
   ///----------
   // -- For robot test shot at interface 5
         L     5;
         T     "DB110_Interf_Program_M1".Program_No_01;

         L     1;
         T     "DB110_Interf_Program_M1".MixingHeadNo;
         L     5;
         T     "DB110_Interf_Program_M1".Robot_01.MC_Place_Number;
         L     201;
         T     "DB110_Interf_Program_M1".Robot_01.Robot_ProgNo_Mould_1;
   ///----------
   // -- For normal interface 5:
   //      L     "DB005_RS<->Extern".MC_Interface[5].FromMC.MouldNumber
   //      T     "DB110_Interf_Program_M1".Program_No_01

   //      L     1
   //      T     "DB110_Interf_Program_M1".MixingHeadNo
   //
   //      L     5
   //      T     "DB110_Interf_Program_M1".Robot_01.MC_Place_Number

   //      L     "DB005_RS<->Extern".MC_Interface[5].FromMC.MouldNumber
   //      T     "DB110_Interf_Program_M1".Robot_01.Robot_ProgNo_Mould_1
         JU    ENDE;
   ///----------
   SS_6: NOP   0;
         AN    "DB110_Interf_Program_M1".Status_IF[6].IF_is_on_1_Position;
         JC    SS_7;
         A     "DB123_MH_IO_Signals".MH[6].IN.MH_Auto_Mode;
         JC    SS6A;
   ///----------
         L     #Temp_ProgNo_MK6_manual;
         L     "DB704_MH_Value".Mixinghead[6].pRrgNumberManual;
         +D;
         T     "DB110_Interf_Program_M1".Program_No_01;
         JU    ENDE;
   ///----------
   SS6A: NOP   0;
         AN    "DB005_RS<->Extern".MC_Interface[6].Data_from_MC.Shot_preperation;
         AN    "DB005_RS<->Extern".MC_Interface[6].Data_from_MC.Shot_release;
         ON    "DB619_State_MPart".SWU[1].SWU_released."06";
         JC    ENDE;
   ///----------
         L     "DB005_RS<->Extern".MC_Interface[6].Data_from_MC.Toolcode;
         T     "DB110_Interf_Program_M1".Program_No_01;

         L     6;
         T     "DB110_Interf_Program_M1".MixingHeadNo;
         T     "DB110_Interf_Program_M1".Robot_01.MC_Place_Number;
         L     "DB005_RS<->Extern".MC_Interface[6].Data_from_MC.Toolcode;
         T     "DB110_Interf_Program_M1".Robot_01.Robot_ProgNo_Mould_1;
         JU    ENDE;

   ///----------
   SS_7: NOP   0;
         AN    "DB110_Interf_Program_M1".Status_IF[7].IF_is_on_1_Position;
         JC    SS_8;
         A     "DB123_MH_IO_Signals".MH[7].IN.MH_Auto_Mode;
         JC    SS7A;
   ///----------
         L     #Temp_ProgNo_MK7_manual;
         L     "DB704_MH_Value".Mixinghead[7].pRrgNumberManual;
         +D;
         T     "DB110_Interf_Program_M1".Program_No_01;
         JU    ENDE;
   ///----------
   SS7A: NOP   0;
         AN    "DB005_RS<->Extern".MC_Interface[7].Data_from_MC.Shot_preperation;
         AN    "DB005_RS<->Extern".MC_Interface[7].Data_from_MC.Shot_release;
         ON    "DB619_State_MPart".SWU[1].SWU_released."07";
         JC    ENDE;
   ///----------
         L     "DB005_RS<->Extern".MC_Interface[7].Data_from_MC.Toolcode;
         T     "DB110_Interf_Program_M1".Program_No_01;

         L     7;
         T     "DB110_Interf_Program_M1".MixingHeadNo;
         T     "DB110_Interf_Program_M1".Robot_01.MC_Place_Number;
         L     "DB005_RS<->Extern".MC_Interface[7].Data_from_MC.Toolcode;
         T     "DB110_Interf_Program_M1".Robot_01.Robot_ProgNo_Mould_1;
         JU    ENDE;

   ///----------
   SS_8: NOP   0;
         AN    "DB110_Interf_Program_M1".Status_IF[8].IF_is_on_1_Position;
         JC    SS_9;
         A     "DB123_MH_IO_Signals".MH[8].IN.MH_Auto_Mode;
         JC    SS8A;
   ///----------
         L     #Temp_ProgNo_MK8_manual;
         L     "DB704_MH_Value".Mixinghead[8].pRrgNumberManual;
         +D;
         T     "DB110_Interf_Program_M1".Program_No_01;
         JU    ENDE;
   ///----------
   SS8A: NOP   0;
         AN    "DB005_RS<->Extern".MC_Interface[8].Data_from_MC.Shot_preperation;
         AN    "DB005_RS<->Extern".MC_Interface[8].Data_from_MC.Shot_release;
         ON    "DB619_State_MPart".SWU[1].SWU_released."08";
         JC    ENDE;
   ///----------
         L     "DB005_RS<->Extern".MC_Interface[8].Data_from_MC.Toolcode;
         T     "DB110_Interf_Program_M1".Program_No_01;

         L     8;
         T     "DB110_Interf_Program_M1".MixingHeadNo;
         T     "DB110_Interf_Program_M1".Robot_01.MC_Place_Number;
         L     "DB005_RS<->Extern".MC_Interface[8].Data_from_MC.Toolcode;
         T     "DB110_Interf_Program_M1".Robot_01.Robot_ProgNo_Mould_1;
         JU    ENDE;
   ///----------
   SS_9: NOP   0;
         AN    "DB110_Interf_Program_M1".Status_IF[9].IF_is_on_1_Position;
         JC    SS_10;
         A     "DB123_MH_IO_Signals".MH[9].IN.MH_Auto_Mode;
         JC    SS9A;
   ///----------
         L     #Temp_ProgNo_MK9_manual;
         L     "DB704_MH_Value".Mixinghead[9].pRrgNumberManual;
         +D;
         T     "DB110_Interf_Program_M1".Program_No_01;
         JU    ENDE;
   ///----------
   SS9A: NOP   0;
         AN    "DB005_RS<->Extern".MC_Interface[9].Data_from_MC.Shot_preperation;
         AN    "DB005_RS<->Extern".MC_Interface[9].Data_from_MC.Shot_release;
         ON    "DB619_State_MPart".SWU[1].SWU_released."09";
         JC    ENDE;
   ///----------
         L     "DB005_RS<->Extern".MC_Interface[9].Data_from_MC.Toolcode;
         T     "DB110_Interf_Program_M1".Program_No_01;

         L     9;
         T     "DB110_Interf_Program_M1".MixingHeadNo;
         T     "DB110_Interf_Program_M1".Robot_01.MC_Place_Number;
         L     "DB005_RS<->Extern".MC_Interface[9].Data_from_MC.Toolcode;
         T     "DB110_Interf_Program_M1".Robot_01.Robot_ProgNo_Mould_1;
         JU    ENDE;
   ///----------
   SS_10:NOP   0;
         AN    "DB110_Interf_Program_M1".Status_IF[10].IF_is_on_1_Position;
         JC    ENDE;
         A     "DB123_MH_IO_Signals".MH[10].IN.MH_Auto_Mode;
         JC    SS10A;
   ///----------
         L     #Temp_ProgNo_MK10_manual;
         L     "DB704_MH_Value".Mixinghead[10].pRrgNumberManual;
         +D;
         T     "DB110_Interf_Program_M1".Program_No_01;
         JU    ENDE;
   ///----------
   SS10A:NOP   0;
         AN    "DB005_RS<->Extern".MC_Interface[10].Data_from_MC.Shot_preperation;
         AN    "DB005_RS<->Extern".MC_Interface[10].Data_from_MC.Shot_release;
         ON    "DB619_State_MPart".SWU[1].SWU_released."10";
         JC    ENDE;
   ///----------
         L     "DB005_RS<->Extern".MC_Interface[10].Data_from_MC.Toolcode;
         T     "DB110_Interf_Program_M1".Program_No_01;

         L     10;
         T     "DB110_Interf_Program_M1".MixingHeadNo;
         T     "DB110_Interf_Program_M1".Robot_01.MC_Place_Number;
         L     "DB005_RS<->Extern".MC_Interface[10].Data_from_MC.Toolcode;
         T     "DB110_Interf_Program_M1".Robot_01.Robot_ProgNo_Mould_1;
         JU    ENDE;
   ///----------
   Test: L     #Temp_ProgNo_MK1_manual;
         T     "DB110_Interf_Program_M1".Program_No_01;
         L     1;
         T     "DB110_Interf_Program_M1".MixingHeadNo;
         JU    ENDE;
   ///----------
   GOON: A     "DB619_State_MPart".Cycle[1].running;
         JC    ENDE;
   ///----------
         L     0;
         T     "DB110_Interf_Program_M1".MixingHeadNo;
   ///---------
         T     "DB110_Interf_Program_M1".Robot_01.MC_Place_Number;
         T     "DB110_Interf_Program_M1".Robot_01.Robot_ProgNo_Mould_1;
         T     "DB110_Interf_Program_M1".Robot_01.Robot_ProgNo_Mould_2;
         T     "DB110_Interf_Program_M1".Robot_01.Robot_ProgNo_Mould_3;
   ///----------
   ENDE: NOP   0;
END_REGION

REGION Network 15: Reset Program number
         AN    "DB619_State_MPart".Cycle[1].running;
         FP    "DB110_Interf_Program_M1".Bits.HF_FP_CycleNotRunning;
         =     "DB110_Interf_Program_M1".Bits.PulseCycleEnd;

         O     "DB110_Interf_Program_M1".Bits.MouldNotReleased;
         O     "DB829_Error_Machine".PouringCycle[1].FLT_WRongStationNumber;
         O     "DB829_Error_Machine".PouringCycle[1].FLT_WrongMixingheadNumber;
         O(;
         O     "DB619_State_MPart".Cycle[1].Pulse_ToolFinished;
         O     "DB110_Interf_Program_M1".Bits.Stop_Cycle;
         O     "DB110_Interf_Program_M1".Bits.PulseCycleEnd;
         AN    "DB829_Error_Machine".PouringCycle[1].FLT_WRongStationNumber;
         AN    "DB829_Error_Machine".PouringCycle[1].FLT_WrongMixingheadNumber;
         );
         FP    "DB110_Interf_Program_M1".Bits.HF_FP_ResetProgramNo;
         JCN   end1;
         L     0;
         T     "DB110_Interf_Program_M1".Program_No_01;
         T     "DB110_Interf_Program_M1".Program_No_02;
   end1: NOP   0;
END_REGION
END_FUNCTION_BLOCK

FUNCTION_BLOCK "FB111_Inerting"   // FB111, STL
{ S7_Optimized_Access := 'FALSE' }
VERSION : 0.1
   VAR_TEMP
      InertPRG : Int;
      dummy : Bool;
      Start_MH : Bool;
      Stop_MH : Bool;
      Purge_On : Bool;
      Purge_Manual : Bool;
      Purge : Bool;
      Inerting : Bool;
      N2_Piston : Bool;
      Shotend : Bool;
      Temp_Release : Bool;
      Shotwight : Real;
      PurgeTime : S5Time;
   END_VAR
BEGIN

REGION Network 1: MH1
         A     "DB123_MH_IO_Signals".MH[1].IN.MH_Manual_Mode;
         JCN   M1Auto;
         L     "DB123_MH_IO_Signals".MH[1].IN.MH_Prog_No_MH;
         T     #InertPRG;

   M1Auto:A     "DB123_MH_IO_Signals".MH[1].IN.MH_Auto_Mode;
         JCN   M1IN;
         L     "DB110_Interf_Program_M1".Signals_ExPlant[1].PrgNo;  // "FRA1>>PrgNr"
         T     #InertPRG;

   M1IN: NOP   0;
         A(;
         A     "DB123_MH_IO_Signals".MH[1].IN.MH_Start;
         A     "DB123_MH_IO_Signals".MH[1].IN.MH_Manual_Mode;
         O;
         A     "DB123_MH_IO_Signals".MH[1].IN.MH_Auto_Mode;
         A(;
         A     "DB005_RS<->Extern".MC_Interface[1].Data_from_MC.Shot_preperation;
         A     "DB704_MH_Value".Mixinghead[1].Conf_IntWithMC;
         O;
         A     "DB110_Interf_Program_M1".Signals_ExPlant[1].Strobe;
         A     "DB704_MH_Value".Mixinghead[1].Conf_IntWithPlantInerface;
         );
         );
         AN    "DB619_State_MPart".Operationmode[1].Test;
         AN    "DB614_MH_State".InertingMH[1].Inert_Off_Dry_Shot;
   //    UN    "DB614_MH_State".InertingMH[2].Inert_runs
   //    UN    "DB614_MH_State".InertingMH[2].OK
   //    UN    "DB614_MH_State".InertingMH[2].Start_PressurizeTimeRuns
         AN    "DB619_State_MPart".Cycle[1].running;
         =     #Start_MH;

